   "Carrier_22_Status.15" AT %I1451.7 : Bool;
   "Carrier_22_SDCFaultCode" AT %IW1452 : Word;   // SDC FAULT CODE
   "Carrier_22_CarrierPosition" AT %ID1454 : DWord;   // CARRIER POSITION
   "Carrier_22_CarrierNumber" AT %IW1458 : Word;   // CARRIER NUMBER
   "Carrier_22_G120DControlWord" AT %IW1460 : Word;   // G120D_STW1_CONTROL
   "Carrier_22_G120DControlWord.0" AT %I1460.0 : Bool;   // Bit_00_ON
   "Carrier_22_G120DControlWord.1" AT %I1460.1 : Bool;   // Bit_01_AUS2_INH
   "Carrier_22_G120DControlWord.2" AT %I1460.2 : Bool;   // Bit_02_AUS3_STOP
   "Carrier_22_G120DControlWord.3" AT %I1460.3 : Bool;   // Bit_03_EN
   "Carrier_22_G120DControlWord.4" AT %I1460.4 : Bool;   // Bit_04_EN_RAMP
   "Carrier_22_G120DControlWord.5" AT %I1460.5 : Bool;   // Bit_05_START_RAMP
   "Carrier_22_G120DControlWord.6" AT %I1460.6 : Bool;   // Bit_06_SETPOINT
   "Carrier_22_G120DControlWord.7" AT %I1460.7 : Bool;   // Bit_07_RESET
   "Carrier_22_G120DControlWord.8" AT %I1461.0 : Bool;   // Bit_08_JOG_R
   "Carrier_22_G120DControlWord.9" AT %I1461.1 : Bool;   // Bit_09_JOG_L
   "Carrier_22_G120DControlWord.10" AT %I1461.2 : Bool;   // Bit_10_CONTR_PLC
   "Carrier_22_G120DControlWord.11" AT %I1461.3 : Bool;   // Bit_11_REVERSE
   "Carrier_22_G120DControlWord.12" AT %I1461.4 : Bool;   // Bit_12_BRAKE_RELEASE
   "Carrier_22_G120DControlWord.13" AT %I1461.5 : Bool;   // Bit_13_DDS
   "Carrier_22_G120DControlWord.14" AT %I1461.6 : Bool;   // Bit_14_DO0
   "Carrier_22_G120DControlWord.15" AT %I1461.7 : Bool;   // Bit_15_DO1
   "Carrier_22_G120DStatusWord" AT %IW1462 : Word;   // G120D_ZSW1_STATUS
   "Carrier_22_G120DStatusWord.0" AT %I1462.0 : Bool;   // Bit_00_READY_RUN
   "Carrier_22_G120DStatusWord.1" AT %I1462.1 : Bool;   // Bit_01_READY_ON
   "Carrier_22_G120DStatusWord.2" AT %I1462.2 : Bool;   // Bit_02_ENABLE
   "Carrier_22_G120DStatusWord.3" AT %I1462.3 : Bool;   // Bit_03_FAULT
   "Carrier_22_G120DStatusWord.4" AT %I1462.4 : Bool;   // Bit_04_OFF2
   "Carrier_22_G120DStatusWord.5" AT %I1462.5 : Bool;   // Bit_05_OFF3
   "Carrier_22_G120DStatusWord.6" AT %I1462.6 : Bool;   // Bit_06_LOCK_OUT
   "Carrier_22_G120DStatusWord.7" AT %I1462.7 : Bool;   // Bit_07_WARN
   "Carrier_22_G120DStatusWord.8" AT %I1463.0 : Bool;   // Bit_08_NO_DEVIATION
   "Carrier_22_G120DStatusWord.9" AT %I1463.1 : Bool;   // Bit_09_CONTR_PLC
   "Carrier_22_G120DStatusWord.10" AT %I1463.2 : Bool;   // Bit_10_F_MAX
   "Carrier_22_G120DStatusWord.11" AT %I1463.3 : Bool;   // Bit_11_LIMIT_REACHED
   "Carrier_22_G120DStatusWord.12" AT %I1463.4 : Bool;   // Bit_12_BRAKE_OPEN
   "Carrier_22_G120DStatusWord.13" AT %I1463.5 : Bool;   // Bit_13_NO_OVERTEMP
   "Carrier_22_G120DStatusWord.14" AT %I1463.6 : Bool;   // Bit_14_CW_CCW
   "Carrier_22_G120DStatusWord.15" AT %I1463.7 : Bool;   // Bit_15_OVERL
   "Carrier_22_Slot2_Input" AT %IW1464 : Word;   // SLOT 2 INPUT WORD
   "Carrier_22_CrashDetectSW" AT %I1464.0 : Bool;   // CRASH DETECT SW
   "Carrier_22_SpareSafetyInput(2_1)" AT %I1464.1 : Bool;   // SPARE SAFETY INPUT
   "Carrier_22_SpareSafetyInput(2_2)" AT %I1464.2 : Bool;   // SPARE SAFETY INPUT
   "Carrier_22_SpareSafetyInput(2_3)" AT %I1464.3 : Bool;   // SPARE SAFETY INPUT
   "Carrier_22_SpareSafetyInput(2_4)" AT %I1464.4 : Bool;   // SPARE SAFETY INPUT
   "Carrier_22_SpareSafetyInput(2_5)" AT %I1464.5 : Bool;   // SPARE SAFETY INPUT
   "Carrier_22_SpareSafetyInput(2_6)" AT %I1464.6 : Bool;   // SPARE SAFETY INPUT
   "Carrier_22_SpareSafetyInput(2_7)" AT %I1464.7 : Bool;   // SPARE SAFETY INPUT
   "Carrier_22_Slot3_SafetyOutput" AT %IW1465 : Word;   // SLOT 3 SAFETY OUTPUT WORD
   "Carrier_22_Crash_Detect_OK" AT %I1465.0 : Bool;   // CARRIER CRASH DETECT
   "Carrier_22_SpareSafetyOutput(3_1)" AT %I1465.1 : Bool;   // SPARE SAFETY OUTPUT
   "Carrier_22_SpareSafetyOutput(3_2)" AT %I1465.2 : Bool;   // SPARE SAFETY OUTPUT
   "Carrier_22_SpareSafetyOutput(3_3)" AT %I1465.3 : Bool;   // SPARE SAFETY OUTPUT
   "Carrier_22_SpareSafetyOutput(3_4)" AT %I1465.4 : Bool;   // SPARE SAFETY OUTPUT
   "Carrier_22_SpareSafetyOutput(3_5)" AT %I1465.5 : Bool;   // SPARE SAFETY OUTPUT
   "Carrier_22_SpareSafetyOutput(3_6)" AT %I1465.6 : Bool;   // SPARE SAFETY OUTPUT
   "Carrier_22_SpareSafetyOutput(3_7)" AT %I1465.7 : Bool;   // SPARE SAFETY OUTPUT
   "Carrier_22_Slot4_Input" AT %IW1466 : Word;   // SLOT 4 INPUT WORD
   "Carrier_22_480VPowerOn_MDCB1" AT %I1466.0 : Bool;   // 480 VAC POWER ON MDCB 1
   "Carrier_22_SpareInput(4_1)" AT %I1466.1 : Bool;   // SPARE INPUT
   "Carrier_22_SpareInput(4_2)" AT %I1466.2 : Bool;   // SPARE INPUT
   "Carrier_22_SitopSelectStatus" AT %I1466.3 : Bool;   // SITOP SELECT STATUS
   "Carrier_22_DCsupplyOnPSCB2" AT %I1466.4 : Bool;   // DC SUPPLY ON PSCB 2
   "Carrier_22_SpareInput(4_5)" AT %I1466.5 : Bool;   // SPARE INPUT
   "Carrier_22_SpareInput(4_6)" AT %I1466.6 : Bool;   // SPARE INPUT
   "Carrier_22_SpareInput(4_7)" AT %I1466.7 : Bool;   // SPARE INPUT
   "Carrier_22_PB1_ProdHoldLH" AT %I1467.0 : Bool;   // PB 1 PRODUCTION HOLD LH
   "Carrier_22_PB2_ResetLH" AT %I1467.1 : Bool;   // PB 2 RESET LH
   "Carrier_22_PB3_ProdHoldRH" AT %I1467.2 : Bool;   // PB 3 PRODUCTION HOLD RH
   "Carrier_22_PB4_ResetRH" AT %I1467.3 : Bool;   // PB 4 RESET RH
   "Carrier_22_SpareInput(4_14)" AT %I1467.4 : Bool;   // SPARE INPUT
   "Carrier_22_SpareInput(4_15)" AT %I1467.5 : Bool;   // SPARE INPUT
   "Carrier_22_SpareInput(4_16)" AT %I1467.6 : Bool;   // SPARE INPUT
   "Carrier_22_SpareInput(4_17)" AT %I1467.7 : Bool;   // SPARE INPUT
   "Carrier_22_Slot5_Output" AT %IW1468 : Word;   // SLOT 5 OUTPUT WORD
   "Carrier_22_IRD400_HMI_24VDC_ENABLE" AT %I1468.0 : Bool;   // IRD 400 PANEL HMI 24V DC POWER
   "Carrier_22_FaultLight_LH" AT %I1468.1 : Bool;   // FAULT LIGHT LH
   "Carrier_22_RunLight_LH" AT %I1468.2 : Bool;   // RUN LIGHT LH
   "Carrier_22_FaultLight_RH" AT %I1468.3 : Bool;   // FAULT LIGHT RH
   "Carrier_22_RunLight_RH" AT %I1468.4 : Bool;   // RUN LIGHT RH
   "Carrier_22_SpareOutput(5_5)" AT %I1468.5 : Bool;   // SPARE OUTPUT
   "Carrier_22_SpareOutput(5_6)" AT %I1468.6 : Bool;   // SPARE OUTPUT
   "Carrier_22_SpareOutput(5_7)" AT %I1468.7 : Bool;   // SPARE OUTPUT
   "Carrier_22_ActualSpeed" AT %IW1470 : Word;   // ACTUAL SPEED
   "Carrier_22_CarrierDriveAlarm" AT %IW1472 : Word;   // CARRIER DRIVE ALARM
   "Carrier_22_CarrierDriveWarning" AT %IW1474 : Word;   // CARRIER DRIVE WARNING
   "Carrier_23_Status" AT %IW1500 : Word;   // CARRIER STATUS WORD
   "Carrier_23_Status.0" AT %I1500.0 : Bool;   // HEARTBEAT
   "Carrier_23_Status.1" AT %I1500.1 : Bool;   // MANUAL
   "Carrier_23_Status.2" AT %I1500.2 : Bool;   // IN_AUTO
   "Carrier_23_Status.3" AT %I1500.3 : Bool;   // POSITIONING_COMPLETE
   "Carrier_23_Status.4" AT %I1500.4 : Bool;   // PRODUCTION HOLD
   "Carrier_23_Status.5" AT %I1500.5 : Bool;   // CARRIER MOVING FORWARD
   "Carrier_23_Status.6" AT %I1500.6 : Bool;   // CARRIER MOVING REVERSE
   "Carrier_23_Status.7" AT %I1500.7 : Bool;   // CARRIER FAULT
   "Carrier_23_Status.8" AT %I1501.0 : Bool;   // CRASH DETECT TRIPPED
   "Carrier_23_Status.9" AT %I1501.1 : Bool;
   "Carrier_23_Status.10" AT %I1501.2 : Bool;
   "Carrier_23_Status.11" AT %I1501.3 : Bool;
   "Carrier_23_Status.12" AT %I1501.4 : Bool;
   "Carrier_23_Status.13" AT %I1501.5 : Bool;
   "Carrier_23_Status.14" AT %I1501.6 : Bool;
   "Carrier_23_Status.15" AT %I1501.7 : Bool;
   "Carrier_23_SDCFaultCode" AT %IW1502 : Word;   // SDC FAULT CODE
   "Carrier_23_CarrierPosition" AT %ID1504 : DWord;   // CARRIER POSITION
   "Carrier_23_CarrierNumber" AT %IW1508 : Word;   // CARRIER NUMBER
   "Carrier_23_G120DControlWord" AT %IW1510 : Word;   // G120D_STW1_CONTROL
   "Carrier_23_G120DControlWord.0" AT %I1510.0 : Bool;   // Bit_00_ON
   "Carrier_23_G120DControlWord.1" AT %I1510.1 : Bool;   // Bit_01_AUS2_INH
   "Carrier_23_G120DControlWord.2" AT %I1510.2 : Bool;   // Bit_02_AUS3_STOP
   "Carrier_23_G120DControlWord.3" AT %I1510.3 : Bool;   // Bit_03_EN
   "Carrier_23_G120DControlWord.4" AT %I1510.4 : Bool;   // Bit_04_EN_RAMP
   "Carrier_23_G120DControlWord.5" AT %I1510.5 : Bool;   // Bit_05_START_RAMP
   "Carrier_23_G120DControlWord.6" AT %I1510.6 : Bool;   // Bit_06_SETPOINT
   "Carrier_23_G120DControlWord.7" AT %I1510.7 : Bool;   // Bit_07_RESET
   "Carrier_23_G120DControlWord.8" AT %I1511.0 : Bool;   // Bit_08_JOG_R
   "Carrier_23_G120DControlWord.9" AT %I1511.1 : Bool;   // Bit_09_JOG_L
   "Carrier_23_G120DControlWord.10" AT %I1511.2 : Bool;   // Bit_10_CONTR_PLC
   "Carrier_23_G120DControlWord.11" AT %I1511.3 : Bool;   // Bit_11_REVERSE
   "Carrier_23_G120DControlWord.12" AT %I1511.4 : Bool;   // Bit_12_BRAKE_RELEASE
   "Carrier_23_G120DControlWord.13" AT %I1511.5 : Bool;   // Bit_13_DDS
   "Carrier_23_G120DControlWord.14" AT %I1511.6 : Bool;   // Bit_14_DO0
   "Carrier_23_G120DControlWord.15" AT %I1511.7 : Bool;   // Bit_15_DO1
   "Carrier_23_G120DStatusWord" AT %IW1512 : Word;   // G120D_ZSW1_STATUS
   "Carrier_23_G120DStatusWord.0" AT %I1512.0 : Bool;   // Bit_00_READY_RUN
   "Carrier_23_G120DStatusWord.1" AT %I1512.1 : Bool;   // Bit_01_READY_ON
   "Carrier_23_G120DStatusWord.2" AT %I1512.2 : Bool;   // Bit_02_ENABLE
   "Carrier_23_G120DStatusWord.3" AT %I1512.3 : Bool;   // Bit_03_FAULT
   "Carrier_23_G120DStatusWord.4" AT %I1512.4 : Bool;   // Bit_04_OFF2
   "Carrier_23_G120DStatusWord.5" AT %I1512.5 : Bool;   // Bit_05_OFF3
   "Carrier_23_G120DStatusWord.6" AT %I1512.6 : Bool;   // Bit_06_LOCK_OUT
   "Carrier_23_G120DStatusWord.7" AT %I1512.7 : Bool;   // Bit_07_WARN
   "Carrier_23_G120DStatusWord.8" AT %I1513.0 : Bool;   // Bit_08_NO_DEVIATION
   "Carrier_23_G120DStatusWord.9" AT %I1513.1 : Bool;   // Bit_09_CONTR_PLC
   "Carrier_23_G120DStatusWord.10" AT %I1513.2 : Bool;   // Bit_10_F_MAX
   "Carrier_23_G120DStatusWord.11" AT %I1513.3 : Bool;   // Bit_11_LIMIT_REACHED
   "Carrier_23_G120DStatusWord.12" AT %I1513.4 : Bool;   // Bit_12_BRAKE_OPEN
   "Carrier_23_G120DStatusWord.13" AT %I1513.5 : Bool;   // Bit_13_NO_OVERTEMP
   "Carrier_23_G120DStatusWord.14" AT %I1513.6 : Bool;   // Bit_14_CW_CCW
   "Carrier_23_G120DStatusWord.15" AT %I1513.7 : Bool;   // Bit_15_OVERL
   "Carrier_23_Slot2_Input" AT %IW1514 : Word;   // SLOT 2 INPUT WORD
   "Carrier_23_CrashDetectSW" AT %I1514.0 : Bool;   // CRASH DETECT SW
   "Carrier_23_SpareSafetyInput(2_1)" AT %I1514.1 : Bool;   // SPARE SAFETY INPUT
   "Carrier_23_SpareSafetyInput(2_2)" AT %I1514.2 : Bool;   // SPARE SAFETY INPUT
   "Carrier_23_SpareSafetyInput(2_3)" AT %I1514.3 : Bool;   // SPARE SAFETY INPUT
   "Carrier_23_SpareSafetyInput(2_4)" AT %I1514.4 : Bool;   // SPARE SAFETY INPUT
   "Carrier_23_SpareSafetyInput(2_5)" AT %I1514.5 : Bool;   // SPARE SAFETY INPUT
   "Carrier_23_SpareSafetyInput(2_6)" AT %I1514.6 : Bool;   // SPARE SAFETY INPUT
   "Carrier_23_SpareSafetyInput(2_7)" AT %I1514.7 : Bool;   // SPARE SAFETY INPUT
   "Carrier_23_Slot3_SafetyOutput" AT %IW1515 : Word;   // SLOT 3 SAFETY OUTPUT WORD
   "Carrier_23_Crash_Detect_OK" AT %I1515.0 : Bool;   // CARRIER CRASH DETECT
   "Carrier_23_SpareSafetyOutput(3_1)" AT %I1515.1 : Bool;   // SPARE SAFETY OUTPUT
   "Carrier_23_SpareSafetyOutput(3_2)" AT %I1515.2 : Bool;   // SPARE SAFETY OUTPUT
   "Carrier_23_SpareSafetyOutput(3_3)" AT %I1515.3 : Bool;   // SPARE SAFETY OUTPUT
   "Carrier_23_SpareSafetyOutput(3_4)" AT %I1515.4 : Bool;   // SPARE SAFETY OUTPUT
   "Carrier_23_SpareSafetyOutput(3_5)" AT %I1515.5 : Bool;   // SPARE SAFETY OUTPUT
   "Carrier_23_SpareSafetyOutput(3_6)" AT %I1515.6 : Bool;   // SPARE SAFETY OUTPUT
   "Carrier_23_SpareSafetyOutput(3_7)" AT %I1515.7 : Bool;   // SPARE SAFETY OUTPUT
   "Carrier_23_Slot4_Input" AT %IW1516 : Word;   // SLOT 4 INPUT WORD
   "Carrier_23_480VPowerOn_MDCB1" AT %I1516.0 : Bool;   // 480 VAC POWER ON MDCB 1
   "Carrier_23_SpareInput(4_1)" AT %I1516.1 : Bool;   // SPARE INPUT
   "Carrier_23_SpareInput(4_2)" AT %I1516.2 : Bool;   // SPARE INPUT
   "Carrier_23_SitopSelectStatus" AT %I1516.3 : Bool;   // SITOP SELECT STATUS
   "Carrier_23_DCsupplyOnPSCB2" AT %I1516.4 : Bool;   // DC SUPPLY ON PSCB 2
   "Carrier_23_SpareInput(4_5)" AT %I1516.5 : Bool;   // SPARE INPUT
   "Carrier_23_SpareInput(4_6)" AT %I1516.6 : Bool;   // SPARE INPUT
   "Carrier_23_SpareInput(4_7)" AT %I1516.7 : Bool;   // SPARE INPUT
   "Carrier_23_PB1_ProdHoldLH" AT %I1517.0 : Bool;   // PB 1 PRODUCTION HOLD LH
   "Carrier_23_PB2_ResetLH" AT %I1517.1 : Bool;   // PB 2 RESET LH
   "Carrier_23_PB3_ProdHoldRH" AT %I1517.2 : Bool;   // PB 3 PRODUCTION HOLD RH
   "Carrier_23_PB4_ResetRH" AT %I1517.3 : Bool;   // PB 4 RESET RH
   "Carrier_23_SpareInput(4_14)" AT %I1517.4 : Bool;   // SPARE INPUT
   "Carrier_23_SpareInput(4_15)" AT %I1517.5 : Bool;   // SPARE INPUT
   "Carrier_23_SpareInput(4_16)" AT %I1517.6 : Bool;   // SPARE INPUT
   "Carrier_23_SpareInput(4_17)" AT %I1517.7 : Bool;   // SPARE INPUT
   "Carrier_23_Slot5_Output" AT %IW1518 : Word;   // SLOT 5 OUTPUT WORD
   "Carrier_23_IRD400_HMI_24VDC_ENABLE" AT %I1518.0 : Bool;   // IRD 400 PANEL HMI 24V DC POWER
   "Carrier_23_FaultLight_LH" AT %I1518.1 : Bool;   // FAULT LIGHT LH
   "Carrier_23_RunLight_LH" AT %I1518.2 : Bool;   // RUN LIGHT LH
   "Carrier_23_FaultLight_RH" AT %I1518.3 : Bool;   // FAULT LIGHT RH
   "Carrier_23_RunLight_RH" AT %I1518.4 : Bool;   // RUN LIGHT RH
   "Carrier_23_SpareOutput(5_5)" AT %I1518.5 : Bool;   // SPARE OUTPUT
   "Carrier_23_SpareOutput(5_6)" AT %I1518.6 : Bool;   // SPARE OUTPUT
   "Carrier_23_SpareOutput(5_7)" AT %I1518.7 : Bool;   // SPARE OUTPUT
   "Carrier_23_ActualSpeed" AT %IW1520 : Word;   // ACTUAL SPEED
   "Carrier_23_CarrierDriveAlarm" AT %IW1522 : Word;   // CARRIER DRIVE ALARM
   "Carrier_23_CarrierDriveWarning" AT %IW1524 : Word;   // CARRIER DRIVE WARNING
   "Carrier_24_Status" AT %IW1550 : Word;   // CARRIER STATUS WORD
   "Carrier_24_Status.0" AT %I1550.0 : Bool;   // HEARTBEAT
   "Carrier_24_Status.1" AT %I1550.1 : Bool;   // MANUAL
   "Carrier_24_Status.2" AT %I1550.2 : Bool;   // IN_AUTO
   "Carrier_24_Status.3" AT %I1550.3 : Bool;   // POSITIONING_COMPLETE
   "Carrier_24_Status.4" AT %I1550.4 : Bool;   // PRODUCTION HOLD
   "Carrier_24_Status.5" AT %I1550.5 : Bool;   // CARRIER MOVING FORWARD
   "Carrier_24_Status.6" AT %I1550.6 : Bool;   // CARRIER MOVING REVERSE
   "Carrier_24_Status.7" AT %I1550.7 : Bool;   // CARRIER FAULT
   "Carrier_24_Status.8" AT %I1551.0 : Bool;   // CRASH DETECT TRIPPED
   "Carrier_24_Status.9" AT %I1551.1 : Bool;
   "Carrier_24_Status.10" AT %I1551.2 : Bool;
   "Carrier_24_Status.11" AT %I1551.3 : Bool;
   "Carrier_24_Status.12" AT %I1551.4 : Bool;
   "Carrier_24_Status.13" AT %I1551.5 : Bool;
   "Carrier_24_Status.14" AT %I1551.6 : Bool;
   "Carrier_24_Status.15" AT %I1551.7 : Bool;
   "Carrier_24_SDCFaultCode" AT %IW1552 : Word;   // SDC FAULT CODE
   "Carrier_24_CarrierPosition" AT %ID1554 : DWord;   // CARRIER POSITION
   "Carrier_24_CarrierNumber" AT %IW1558 : Word;   // CARRIER NUMBER
   "Carrier_24_G120DControlWord" AT %IW1560 : Word;   // G120D_STW1_CONTROL
   "Carrier_24_G120DControlWord.0" AT %I1560.0 : Bool;   // Bit_00_ON
   "Carrier_24_G120DControlWord.1" AT %I1560.1 : Bool;   // Bit_01_AUS2_INH
   "Carrier_24_G120DControlWord.2" AT %I1560.2 : Bool;   // Bit_02_AUS3_STOP
   "Carrier_24_G120DControlWord.3" AT %I1560.3 : Bool;   // Bit_03_EN
   "Carrier_24_G120DControlWord.4" AT %I1560.4 : Bool;   // Bit_04_EN_RAMP
   "Carrier_24_G120DControlWord.5" AT %I1560.5 : Bool;   // Bit_05_START_RAMP
   "Carrier_24_G120DControlWord.6" AT %I1560.6 : Bool;   // Bit_06_SETPOINT
   "Carrier_24_G120DControlWord.7" AT %I1560.7 : Bool;   // Bit_07_RESET
   "Carrier_24_G120DControlWord.8" AT %I1561.0 : Bool;   // Bit_08_JOG_R
   "Carrier_24_G120DControlWord.9" AT %I1561.1 : Bool;   // Bit_09_JOG_L
   "Carrier_24_G120DControlWord.10" AT %I1561.2 : Bool;   // Bit_10_CONTR_PLC
   "Carrier_24_G120DControlWord.11" AT %I1561.3 : Bool;   // Bit_11_REVERSE
   "Carrier_24_G120DControlWord.12" AT %I1561.4 : Bool;   // Bit_12_BRAKE_RELEASE
   "Carrier_24_G120DControlWord.13" AT %I1561.5 : Bool;   // Bit_13_DDS
   "Carrier_24_G120DControlWord.14" AT %I1561.6 : Bool;   // Bit_14_DO0
   "Carrier_24_G120DControlWord.15" AT %I1561.7 : Bool;   // Bit_15_DO1
   "Carrier_24_G120DStatusWord" AT %IW1562 : Word;   // G120D_ZSW1_STATUS
   "Carrier_24_G120DStatusWord.0" AT %I1562.0 : Bool;   // Bit_00_READY_RUN
   "Carrier_24_G120DStatusWord.1" AT %I1562.1 : Bool;   // Bit_01_READY_ON
   "Carrier_24_G120DStatusWord.2" AT %I1562.2 : Bool;   // Bit_02_ENABLE
   "Carrier_24_G120DStatusWord.3" AT %I1562.3 : Bool;   // Bit_03_FAULT
   "Carrier_24_G120DStatusWord.4" AT %I1562.4 : Bool;   // Bit_04_OFF2
   "Carrier_24_G120DStatusWord.5" AT %I1562.5 : Bool;   // Bit_05_OFF3
   "Carrier_24_G120DStatusWord.6" AT %I1562.6 : Bool;   // Bit_06_LOCK_OUT
   "Carrier_24_G120DStatusWord.7" AT %I1562.7 : Bool;   // Bit_07_WARN
   "Carrier_24_G120DStatusWord.8" AT %I1563.0 : Bool;   // Bit_08_NO_DEVIATION
   "Carrier_24_G120DStatusWord.9" AT %I1563.1 : Bool;   // Bit_09_CONTR_PLC
   "Carrier_24_G120DStatusWord.10" AT %I1563.2 : Bool;   // Bit_10_F_MAX
   "Carrier_24_G120DStatusWord.11" AT %I1563.3 : Bool;   // Bit_11_LIMIT_REACHED
   "Carrier_24_G120DStatusWord.12" AT %I1563.4 : Bool;   // Bit_12_BRAKE_OPEN
   "Carrier_24_G120DStatusWord.13" AT %I1563.5 : Bool;   // Bit_13_NO_OVERTEMP
   "Carrier_24_G120DStatusWord.14" AT %I1563.6 : Bool;   // Bit_14_CW_CCW
   "Carrier_24_G120DStatusWord.15" AT %I1563.7 : Bool;   // Bit_15_OVERL
   "Carrier_24_Slot2_Input" AT %IW1564 : Word;   // SLOT 2 INPUT WORD
   "Carrier_24_CrashDetectSW" AT %I1564.0 : Bool;   // CRASH DETECT SW
   "Carrier_24_SpareSafetyInput(2_1)" AT %I1564.1 : Bool;   // SPARE SAFETY INPUT
   "Carrier_24_SpareSafetyInput(2_2)" AT %I1564.2 : Bool;   // SPARE SAFETY INPUT
   "Carrier_24_SpareSafetyInput(2_3)" AT %I1564.3 : Bool;   // SPARE SAFETY INPUT
   "Carrier_24_SpareSafetyInput(2_4)" AT %I1564.4 : Bool;   // SPARE SAFETY INPUT
   "Carrier_24_SpareSafetyInput(2_5)" AT %I1564.5 : Bool;   // SPARE SAFETY INPUT
   "Carrier_24_SpareSafetyInput(2_6)" AT %I1564.6 : Bool;   // SPARE SAFETY INPUT
   "Carrier_24_SpareSafetyInput(2_7)" AT %I1564.7 : Bool;   // SPARE SAFETY INPUT
   "Carrier_24_Slot3_SafetyOutput" AT %IW1565 : Word;   // SLOT 3 SAFETY OUTPUT WORD
   "Carrier_24_Crash_Detect_OK" AT %I1565.0 : Bool;   // CARRIER CRASH DETECT
   "Carrier_24_SpareSafetyOutput(3_1)" AT %I1565.1 : Bool;   // SPARE SAFETY OUTPUT
   "Carrier_24_SpareSafetyOutput(3_2)" AT %I1565.2 : Bool;   // SPARE SAFETY OUTPUT
   "Carrier_24_SpareSafetyOutput(3_3)" AT %I1565.3 : Bool;   // SPARE SAFETY OUTPUT
   "Carrier_24_SpareSafetyOutput(3_4)" AT %I1565.4 : Bool;   // SPARE SAFETY OUTPUT
   "Carrier_24_SpareSafetyOutput(3_5)" AT %I1565.5 : Bool;   // SPARE SAFETY OUTPUT
   "Carrier_24_SpareSafetyOutput(3_6)" AT %I1565.6 : Bool;   // SPARE SAFETY OUTPUT
   "Carrier_24_SpareSafetyOutput(3_7)" AT %I1565.7 : Bool;   // SPARE SAFETY OUTPUT
   "Carrier_24_Slot4_Input" AT %IW1566 : Word;   // SLOT 4 INPUT WORD
   "Carrier_24_480VPowerOn_MDCB1" AT %I1566.0 : Bool;   // 480 VAC POWER ON MDCB 1
   "Carrier_24_SpareInput(4_1)" AT %I1566.1 : Bool;   // SPARE INPUT
   "Carrier_24_SpareInput(4_2)" AT %I1566.2 : Bool;   // SPARE INPUT
   "Carrier_24_SitopSelectStatus" AT %I1566.3 : Bool;   // SITOP SELECT STATUS
   "Carrier_24_DCsupplyOnPSCB2" AT %I1566.4 : Bool;   // DC SUPPLY ON PSCB 2
   "Carrier_24_SpareInput(4_5)" AT %I1566.5 : Bool;   // SPARE INPUT
   "Carrier_24_SpareInput(4_6)" AT %I1566.6 : Bool;   // SPARE INPUT
   "Carrier_24_SpareInput(4_7)" AT %I1566.7 : Bool;   // SPARE INPUT
   "Carrier_24_PB1_ProdHoldLH" AT %I1567.0 : Bool;   // PB 1 PRODUCTION HOLD LH
   "Carrier_24_PB2_ResetLH" AT %I1567.1 : Bool;   // PB 2 RESET LH
   "Carrier_24_PB3_ProdHoldRH" AT %I1567.2 : Bool;   // PB 3 PRODUCTION HOLD RH
   "Carrier_24_PB4_ResetRH" AT %I1567.3 : Bool;   // PB 4 RESET RH
   "Carrier_24_SpareInput(4_14)" AT %I1567.4 : Bool;   // SPARE INPUT
   "Carrier_24_SpareInput(4_15)" AT %I1567.5 : Bool;   // SPARE INPUT
   "Carrier_24_SpareInput(4_16)" AT %I1567.6 : Bool;   // SPARE INPUT
   "Carrier_24_SpareInput(4_17)" AT %I1567.7 : Bool;   // SPARE INPUT
   "Carrier_24_Slot5_Output" AT %IW1568 : Word;   // SLOT 5 OUTPUT WORD
   "Carrier_24_IRD400_HMI_24VDC_ENABLE" AT %I1568.0 : Bool;   // IRD 400 PANEL HMI 24V DC POWER
   "Carrier_24_FaultLight_LH" AT %I1568.1 : Bool;   // FAULT LIGHT LH
   "Carrier_24_RunLight_LH" AT %I1568.2 : Bool;   // RUN LIGHT LH
   "Carrier_24_FaultLight_RH" AT %I1568.3 : Bool;   // FAULT LIGHT RH
   "Carrier_24_RunLight_RH" AT %I1568.4 : Bool;   // RUN LIGHT RH
   "Carrier_24_SpareOutput(5_5)" AT %I1568.5 : Bool;   // SPARE OUTPUT
   "Carrier_24_SpareOutput(5_6)" AT %I1568.6 : Bool;   // SPARE OUTPUT
   "Carrier_24_SpareOutput(5_7)" AT %I1568.7 : Bool;   // SPARE OUTPUT
   "Carrier_24_ActualSpeed" AT %IW1570 : Word;   // ACTUAL SPEED
   "Carrier_24_CarrierDriveAlarm" AT %IW1572 : Word;   // CARRIER DRIVE ALARM
   "Carrier_24_CarrierDriveWarning" AT %IW1574 : Word;   // CARRIER DRIVE WARNING
   "Carrier_25_Status" AT %IW1600 : Word;   // CARRIER STATUS WORD
   "Carrier_25_Status.0" AT %I1600.0 : Bool;   // HEARTBEAT
   "Carrier_25_Status.1" AT %I1600.1 : Bool;   // MANUAL
   "Carrier_25_Status.2" AT %I1600.2 : Bool;   // IN_AUTO
   "Carrier_25_Status.3" AT %I1600.3 : Bool;   // POSITIONING_COMPLETE
   "Carrier_25_Status.4" AT %I1600.4 : Bool;   // PRODUCTION HOLD
   "Carrier_25_Status.5" AT %I1600.5 : Bool;   // CARRIER MOVING FORWARD
   "Carrier_25_Status.6" AT %I1600.6 : Bool;   // CARRIER MOVING REVERSE
   "Carrier_25_Status.7" AT %I1600.7 : Bool;   // CARRIER FAULT
   "Carrier_25_Status.8" AT %I1601.0 : Bool;   // CRASH DETECT TRIPPED
   "Carrier_25_Status.9" AT %I1601.1 : Bool;
   "Carrier_25_Status.10" AT %I1601.2 : Bool;
   "Carrier_25_Status.11" AT %I1601.3 : Bool;
   "Carrier_25_Status.12" AT %I1601.4 : Bool;
   "Carrier_25_Status.13" AT %I1601.5 : Bool;
   "Carrier_25_Status.14" AT %I1601.6 : Bool;
   "Carrier_25_Status.15" AT %I1601.7 : Bool;
   "Carrier_25_SDCFaultCode" AT %IW1602 : Word;   // SDC FAULT CODE
   "Carrier_25_CarrierPosition" AT %ID1604 : DWord;   // CARRIER POSITION
   "Carrier_25_CarrierNumber" AT %IW1608 : Word;   // CARRIER NUMBER
   "Carrier_25_G120DControlWord" AT %IW1610 : Word;   // G120D_STW1_CONTROL
   "Carrier_25_G120DControlWord.0" AT %I1610.0 : Bool;   // Bit_00_ON
   "Carrier_25_G120DControlWord.1" AT %I1610.1 : Bool;   // Bit_01_AUS2_INH
   "Carrier_25_G120DControlWord.2" AT %I1610.2 : Bool;   // Bit_02_AUS3_STOP
   "Carrier_25_G120DControlWord.3" AT %I1610.3 : Bool;   // Bit_03_EN
   "Carrier_25_G120DControlWord.4" AT %I1610.4 : Bool;   // Bit_04_EN_RAMP
   "Carrier_25_G120DControlWord.5" AT %I1610.5 : Bool;   // Bit_05_START_RAMP
   "Carrier_25_G120DControlWord.6" AT %I1610.6 : Bool;   // Bit_06_SETPOINT
   "Carrier_25_G120DControlWord.7" AT %I1610.7 : Bool;   // Bit_07_RESET
   "Carrier_25_G120DControlWord.8" AT %I1611.0 : Bool;   // Bit_08_JOG_R
   "Carrier_25_G120DControlWord.9" AT %I1611.1 : Bool;   // Bit_09_JOG_L
   "Carrier_25_G120DControlWord.10" AT %I1611.2 : Bool;   // Bit_10_CONTR_PLC
   "Carrier_25_G120DControlWord.11" AT %I1611.3 : Bool;   // Bit_11_REVERSE
   "Carrier_25_G120DControlWord.12" AT %I1611.4 : Bool;   // Bit_12_BRAKE_RELEASE
   "Carrier_25_G120DControlWord.13" AT %I1611.5 : Bool;   // Bit_13_DDS
   "Carrier_25_G120DControlWord.14" AT %I1611.6 : Bool;   // Bit_14_DO0
   "Carrier_25_G120DControlWord.15" AT %I1611.7 : Bool;   // Bit_15_DO1
   "Carrier_25_G120DStatusWord" AT %IW1612 : Word;   // G120D_ZSW1_STATUS
   "Carrier_25_G120DStatusWord.0" AT %I1612.0 : Bool;   // Bit_00_READY_RUN
   "Carrier_25_G120DStatusWord.1" AT %I1612.1 : Bool;   // Bit_01_READY_ON
   "Carrier_25_G120DStatusWord.2" AT %I1612.2 : Bool;   // Bit_02_ENABLE
   "Carrier_25_G120DStatusWord.3" AT %I1612.3 : Bool;   // Bit_03_FAULT
   "Carrier_25_G120DStatusWord.4" AT %I1612.4 : Bool;   // Bit_04_OFF2
   "Carrier_25_G120DStatusWord.5" AT %I1612.5 : Bool;   // Bit_05_OFF3
   "Carrier_25_G120DStatusWord.6" AT %I1612.6 : Bool;   // Bit_06_LOCK_OUT
   "Carrier_25_G120DStatusWord.7" AT %I1612.7 : Bool;   // Bit_07_WARN
   "Carrier_25_G120DStatusWord.8" AT %I1613.0 : Bool;   // Bit_08_NO_DEVIATION
   "Carrier_25_G120DStatusWord.9" AT %I1613.1 : Bool;   // Bit_09_CONTR_PLC
   "Carrier_25_G120DStatusWord.10" AT %I1613.2 : Bool;   // Bit_10_F_MAX
   "Carrier_25_G120DStatusWord.11" AT %I1613.3 : Bool;   // Bit_11_LIMIT_REACHED
   "Carrier_25_G120DStatusWord.12" AT %I1613.4 : Bool;   // Bit_12_BRAKE_OPEN
   "Carrier_25_G120DStatusWord.13" AT %I1613.5 : Bool;   // Bit_13_NO_OVERTEMP
   "Carrier_25_G120DStatusWord.14" AT %I1613.6 : Bool;   // Bit_14_CW_CCW
   "Carrier_25_G120DStatusWord.15" AT %I1613.7 : Bool;   // Bit_15_OVERL
   "Carrier_25_Slot2_Input" AT %IW1614 : Word;   // SLOT 2 INPUT WORD
   "Carrier_25_CrashDetectSW" AT %I1614.0 : Bool;   // CRASH DETECT SW
   "Carrier_25_SpareSafetyInput(2_1)" AT %I1614.1 : Bool;   // SPARE SAFETY INPUT
   "Carrier_25_SpareSafetyInput(2_2)" AT %I1614.2 : Bool;   // SPARE SAFETY INPUT
   "Carrier_25_SpareSafetyInput(2_3)" AT %I1614.3 : Bool;   // SPARE SAFETY INPUT
   "Carrier_25_SpareSafetyInput(2_4)" AT %I1614.4 : Bool;   // SPARE SAFETY INPUT
   "Carrier_25_SpareSafetyInput(2_5)" AT %I1614.5 : Bool;   // SPARE SAFETY INPUT
   "Carrier_25_SpareSafetyInput(2_6)" AT %I1614.6 : Bool;   // SPARE SAFETY INPUT
   "Carrier_25_SpareSafetyInput(2_7)" AT %I1614.7 : Bool;   // SPARE SAFETY INPUT
   "Carrier_25_Slot3_SafetyOutput" AT %IW1615 : Word;   // SLOT 3 SAFETY OUTPUT WORD
   "Carrier_25_Crash_Detect_OK" AT %I1615.0 : Bool;   // CARRIER CRASH DETECT
   "Carrier_25_SpareSafetyOutput(3_1)" AT %I1615.1 : Bool;   // SPARE SAFETY OUTPUT
   "Carrier_25_SpareSafetyOutput(3_2)" AT %I1615.2 : Bool;   // SPARE SAFETY OUTPUT
   "Carrier_25_SpareSafetyOutput(3_3)" AT %I1615.3 : Bool;   // SPARE SAFETY OUTPUT
   "Carrier_25_SpareSafetyOutput(3_4)" AT %I1615.4 : Bool;   // SPARE SAFETY OUTPUT
   "Carrier_25_SpareSafetyOutput(3_5)" AT %I1615.5 : Bool;   // SPARE SAFETY OUTPUT
   "Carrier_25_SpareSafetyOutput(3_6)" AT %I1615.6 : Bool;   // SPARE SAFETY OUTPUT
   "Carrier_25_SpareSafetyOutput(3_7)" AT %I1615.7 : Bool;   // SPARE SAFETY OUTPUT
   "Carrier_25_Slot4_Input" AT %IW1616 : Word;   // SLOT 4 INPUT WORD
   "Carrier_25_480VPowerOn_MDCB1" AT %I1616.0 : Bool;   // 480 VAC POWER ON MDCB 1
   "Carrier_25_SpareInput(4_1)" AT %I1616.1 : Bool;   // SPARE INPUT
   "Carrier_25_SpareInput(4_2)" AT %I1616.2 : Bool;   // SPARE INPUT
   "Carrier_25_SitopSelectStatus" AT %I1616.3 : Bool;   // SITOP SELECT STATUS
   "Carrier_25_DCsupplyOnPSCB2" AT %I1616.4 : Bool;   // DC SUPPLY ON PSCB 2
   "Carrier_25_SpareInput(4_5)" AT %I1616.5 : Bool;   // SPARE INPUT
   "Carrier_25_SpareInput(4_6)" AT %I1616.6 : Bool;   // SPARE INPUT
   "Carrier_25_SpareInput(4_7)" AT %I1616.7 : Bool;   // SPARE INPUT
   "Carrier_25_PB1_ProdHoldLH" AT %I1617.0 : Bool;   // PB 1 PRODUCTION HOLD LH
   "Carrier_25_PB2_ResetLH" AT %I1617.1 : Bool;   // PB 2 RESET LH
   "Carrier_25_PB3_ProdHoldRH" AT %I1617.2 : Bool;   // PB 3 PRODUCTION HOLD RH
   "Carrier_25_PB4_ResetRH" AT %I1617.3 : Bool;   // PB 4 RESET RH
   "Carrier_25_SpareInput(4_14)" AT %I1617.4 : Bool;   // SPARE INPUT
   "Carrier_25_SpareInput(4_15)" AT %I1617.5 : Bool;   // SPARE INPUT
   "Carrier_25_SpareInput(4_16)" AT %I1617.6 : Bool;   // SPARE INPUT
   "Carrier_25_SpareInput(4_17)" AT %I1617.7 : Bool;   // SPARE INPUT
   "Carrier_25_Slot5_Output" AT %IW1618 : Word;   // SLOT 5 OUTPUT WORD
   "Carrier_25_IRD400_HMI_24VDC_ENABLE" AT %I1618.0 : Bool;   // IRD 400 PANEL HMI 24V DC POWER
   "Carrier_25_FaultLight_LH" AT %I1618.1 : Bool;   // FAULT LIGHT LH
   "Carrier_25_RunLight_LH" AT %I1618.2 : Bool;   // RUN LIGHT LH
   "Carrier_25_FaultLight_RH" AT %I1618.3 : Bool;   // FAULT LIGHT RH
   "Carrier_25_RunLight_RH" AT %I1618.4 : Bool;   // RUN LIGHT RH
   "Carrier_25_SpareOutput(5_5)" AT %I1618.5 : Bool;   // SPARE OUTPUT
   "Carrier_25_SpareOutput(5_6)" AT %I1618.6 : Bool;   // SPARE OUTPUT
   "Carrier_25_SpareOutput(5_7)" AT %I1618.7 : Bool;   // SPARE OUTPUT
   "Carrier_25_ActualSpeed" AT %IW1620 : Word;   // ACTUAL SPEED
   "Carrier_25_CarrierDriveAlarm" AT %IW1622 : Word;   // CARRIER DRIVE ALARM
   "Carrier_25_CarrierDriveWarning" AT %IW1624 : Word;   // CARRIER DRIVE WARNING
   "Carrier_26_Status" AT %IW1650 : Word;   // CARRIER STATUS WORD
   "Carrier_26_Status.0" AT %I1650.0 : Bool;   // HEARTBEAT
   "Carrier_26_Status.1" AT %I1650.1 : Bool;   // MANUAL
   "Carrier_26_Status.2" AT %I1650.2 : Bool;   // IN_AUTO
   "Carrier_26_Status.3" AT %I1650.3 : Bool;   // POSITIONING_COMPLETE
   "Carrier_26_Status.4" AT %I1650.4 : Bool;   // PRODUCTION HOLD
   "Carrier_26_Status.5" AT %I1650.5 : Bool;   // CARRIER MOVING FORWARD
   "Carrier_26_Status.6" AT %I1650.6 : Bool;   // CARRIER MOVING REVERSE
   "Carrier_26_Status.7" AT %I1650.7 : Bool;   // CARRIER FAULT
   "Carrier_26_Status.8" AT %I1651.0 : Bool;   // CRASH DETECT TRIPPED
   "Carrier_26_Status.9" AT %I1651.1 : Bool;
   "Carrier_26_Status.10" AT %I1651.2 : Bool;
   "Carrier_26_Status.11" AT %I1651.3 : Bool;
   "Carrier_26_Status.12" AT %I1651.4 : Bool;
   "Carrier_26_Status.13" AT %I1651.5 : Bool;
   "Carrier_26_Status.14" AT %I1651.6 : Bool;
   "Carrier_26_Status.15" AT %I1651.7 : Bool;
   "Carrier_26_SDCFaultCode" AT %IW1652 : Word;   // SDC FAULT CODE
   "Carrier_26_CarrierPosition" AT %ID1654 : DWord;   // CARRIER POSITION
   "Carrier_26_CarrierNumber" AT %IW1658 : Word;   // CARRIER NUMBER
   "Carrier_26_G120DControlWord" AT %IW1660 : Word;   // G120D_STW1_CONTROL
   "Carrier_26_G120DControlWord.0" AT %I1660.0 : Bool;   // Bit_00_ON
   "Carrier_26_G120DControlWord.1" AT %I1660.1 : Bool;   // Bit_01_AUS2_INH
   "Carrier_26_G120DControlWord.2" AT %I1660.2 : Bool;   // Bit_02_AUS3_STOP
   "Carrier_26_G120DControlWord.3" AT %I1660.3 : Bool;   // Bit_03_EN
   "Carrier_26_G120DControlWord.4" AT %I1660.4 : Bool;   // Bit_04_EN_RAMP
   "Carrier_26_G120DControlWord.5" AT %I1660.5 : Bool;   // Bit_05_START_RAMP
   "Carrier_26_G120DControlWord.6" AT %I1660.6 : Bool;   // Bit_06_SETPOINT
   "Carrier_26_G120DControlWord.7" AT %I1660.7 : Bool;   // Bit_07_RESET
   "Carrier_26_G120DControlWord.8" AT %I1661.0 : Bool;   // Bit_08_JOG_R
   "Carrier_26_G120DControlWord.9" AT %I1661.1 : Bool;   // Bit_09_JOG_L
   "Carrier_26_G120DControlWord.10" AT %I1661.2 : Bool;   // Bit_10_CONTR_PLC
   "Carrier_26_G120DControlWord.11" AT %I1661.3 : Bool;   // Bit_11_REVERSE
   "Carrier_26_G120DControlWord.12" AT %I1661.4 : Bool;   // Bit_12_BRAKE_RELEASE
   "Carrier_26_G120DControlWord.13" AT %I1661.5 : Bool;   // Bit_13_DDS
   "Carrier_26_G120DControlWord.14" AT %I1661.6 : Bool;   // Bit_14_DO0
   "Carrier_26_G120DControlWord.15" AT %I1661.7 : Bool;   // Bit_15_DO1
   "Carrier_26_G120DStatusWord" AT %IW1662 : Word;   // G120D_ZSW1_STATUS
   "Carrier_26_G120DStatusWord.0" AT %I1662.0 : Bool;   // Bit_00_READY_RUN
   "Carrier_26_G120DStatusWord.1" AT %I1662.1 : Bool;   // Bit_01_READY_ON
   "Carrier_26_G120DStatusWord.2" AT %I1662.2 : Bool;   // Bit_02_ENABLE
   "Carrier_26_G120DStatusWord.3" AT %I1662.3 : Bool;   // Bit_03_FAULT
   "Carrier_26_G120DStatusWord.4" AT %I1662.4 : Bool;   // Bit_04_OFF2
   "Carrier_26_G120DStatusWord.5" AT %I1662.5 : Bool;   // Bit_05_OFF3
   "Carrier_26_G120DStatusWord.6" AT %I1662.6 : Bool;   // Bit_06_LOCK_OUT
   "Carrier_26_G120DStatusWord.7" AT %I1662.7 : Bool;   // Bit_07_WARN
   "Carrier_26_G120DStatusWord.8" AT %I1663.0 : Bool;   // Bit_08_NO_DEVIATION
   "Carrier_26_G120DStatusWord.9" AT %I1663.1 : Bool;   // Bit_09_CONTR_PLC
   "Carrier_26_G120DStatusWord.10" AT %I1663.2 : Bool;   // Bit_10_F_MAX
   "Carrier_26_G120DStatusWord.11" AT %I1663.3 : Bool;   // Bit_11_LIMIT_REACHED
   "Carrier_26_G120DStatusWord.12" AT %I1663.4 : Bool;   // Bit_12_BRAKE_OPEN
   "Carrier_26_G120DStatusWord.13" AT %I1663.5 : Bool;   // Bit_13_NO_OVERTEMP
   "Carrier_26_G120DStatusWord.14" AT %I1663.6 : Bool;   // Bit_14_CW_CCW
   "Carrier_26_G120DStatusWord.15" AT %I1663.7 : Bool;   // Bit_15_OVERL
   "Carrier_26_Slot2_Input" AT %IW1664 : Word;   // SLOT 2 INPUT WORD
   "Carrier_26_CrashDetectSW" AT %I1664.0 : Bool;   // CRASH DETECT SW
   "Carrier_26_SpareSafetyInput(2_1)" AT %I1664.1 : Bool;   // SPARE SAFETY INPUT
   "Carrier_26_SpareSafetyInput(2_2)" AT %I1664.2 : Bool;   // SPARE SAFETY INPUT
   "Carrier_26_SpareSafetyInput(2_3)" AT %I1664.3 : Bool;   // SPARE SAFETY INPUT
   "Carrier_26_SpareSafetyInput(2_4)" AT %I1664.4 : Bool;   // SPARE SAFETY INPUT
   "Carrier_26_SpareSafetyInput(2_5)" AT %I1664.5 : Bool;   // SPARE SAFETY INPUT
   "Carrier_26_SpareSafetyInput(2_6)" AT %I1664.6 : Bool;   // SPARE SAFETY INPUT
   "Carrier_26_SpareSafetyInput(2_7)" AT %I1664.7 : Bool;   // SPARE SAFETY INPUT
   "Carrier_26_Slot3_SafetyOutput" AT %IW1665 : Word;   // SLOT 3 SAFETY OUTPUT WORD
   "Carrier_26_Crash_Detect_OK" AT %I1665.0 : Bool;   // CARRIER CRASH DETECT
   "Carrier_26_SpareSafetyOutput(3_1)" AT %I1665.1 : Bool;   // SPARE SAFETY OUTPUT
   "Carrier_26_SpareSafetyOutput(3_2)" AT %I1665.2 : Bool;   // SPARE SAFETY OUTPUT
   "Carrier_26_SpareSafetyOutput(3_3)" AT %I1665.3 : Bool;   // SPARE SAFETY OUTPUT
   "Carrier_26_SpareSafetyOutput(3_4)" AT %I1665.4 : Bool;   // SPARE SAFETY OUTPUT
   "Carrier_26_SpareSafetyOutput(3_5)" AT %I1665.5 : Bool;   // SPARE SAFETY OUTPUT
